// TIA Portal project "EbAndon v2_0_1" (V15) (continued)
TYPE "Color Library"
   STRUCT
      BkBk : USInt := 0;
      BgWh : USInt := 1;
      FgWh : USInt := 2;
      FlWh : USInt := 3;
      BgGray : USInt := 4;
      FgGray : USInt := 5;
      FlGray : USInt := 6;
      BgLRd : USInt := 7;
      FgLRd : USInt := 8;
      FlLRd : USInt := 9;
      BgDRd : USInt := 10;
      FgDRd : USInt := 11;
      FlDrd : USInt := 12;
      BgLYe : USInt := 13;
      FgLYe : USInt := 14;
      FlLYe : USInt := 15;
      BgDYe : USInt := 16;
      FgDYe : USInt := 17;
      FlDYe : USInt := 18;
      BgLGr : USInt := 19;
      FgLGr : USInt := 20;
      FlLGr : USInt := 21;
      BgDGr : USInt := 22;
      FgDGr : USInt := 23;
      FlDGr : USInt := 24;
      BgLTe : USInt := 25;
      FgLTe : USInt := 26;
      FlLTe : USInt := 27;
      BgDTe : USInt := 28;
      FgDTe : USInt := 29;
      FlDTe : USInt := 30;
      BgLBl : USInt := 31;
      FgLBl : USInt := 32;
      FlLBl : USInt := 33;
      BgDBl : USInt := 34;
      FgDBl : USInt := 35;
      FlDBl : USInt := 36;
      BgLPu : USInt := 37;
      FgLPu : USInt := 38;
      FlLPu : USInt := 39;
      BgDPu : USInt := 40;
      FgDPu : USInt := 41;
      FlDPu : USInt := 42;
      disabled : USInt := 254;
      invisible : USInt := 255;
   END_STRUCT;
END_TYPE

TYPE "Station Assignment: Button Details"
   STRUCT
      alloted : Struct
         animate : USInt;
         value : WString[10];
      END_STRUCT;
      critical : Struct
         animate : USInt;
         value : WString[10];
      END_STRUCT;
      label : Struct
         animate : USInt;
         value : WString[2];
      END_STRUCT;
      partNumber : Struct
         animate : USInt;
         value : WString[40];
      END_STRUCT;
      select : Struct
         actuate : Bool;
         animate : USInt;
      END_STRUCT;
   END_STRUCT;
END_TYPE

TYPE "IO Field Data: Part Number"
   STRUCT
      animate : USInt;
      inputFinished : Bool;
      value : WString[40];
   END_STRUCT;
END_TYPE

TYPE "Line Label Data"
   STRUCT
      animate : Struct
         bg : USInt;
         ioField : USInt;
      END_STRUCT;
      inputFinished : Bool;
      value : WString[10];
   END_STRUCT;
END_TYPE

TYPE "Drop Zone Data"
   STRUCT
      animate : Struct
         bg : USInt;
         ioField : USInt;
      END_STRUCT;
      inputFinished : Bool;
      value : WString[10];
   END_STRUCT;
END_TYPE

TYPE "IO Field Data: Timers"
   STRUCT
      animate : USInt;
      inputFinished : Bool;
      value : WString[5];
   END_STRUCT;
END_TYPE

TYPE "Table Nav"
   STRUCT
      top : "PB Data: Graphic/Text List";
      pageUp : "PB Data: Graphic/Text List";
      lineUp : "PB Data: Graphic/Text List";
      lineDown : "PB Data: Graphic/Text List";
      pageDown : "PB Data: Graphic/Text List";
      bottom : "PB Data: Graphic/Text List";
   END_STRUCT;
END_TYPE

DATA_BLOCK "EMP IDB"   // DB1
{ S7_Optimized_Access := 'TRUE' }
VERSION : 0.1
// stored: InstanceOfName EMP
"EMP"
BEGIN
   constants.buttonCount := 8;
   stations.current[0].presetTime.allotted[7] := 1800.0;
   stations.current[0].presetTime.allotted[3] := 1800.0;
   stations.current[0].presetTime.critical[7] := 300.0;
   stations.current[0].presetTime.critical[3] := 300.0;
   stations.current[0].partNumbers[7] := WSTRING#'16.32.112.500.100A';
   stations.current[0].partNumbers[6] := WSTRING#'';
   stations.current[0].partNumbers[5] := WSTRING#'';
   stations.current[0].partNumbers[3] := WSTRING#'16.32.112.500.220A';
   stations.current[0].partNumbers[2] := WSTRING#'';
   stations.current[0].partNumbers[1] := WSTRING#'';
   stations.current[0].line := WSTRING#'VOLVO 16';
   stations.current[1].line := WSTRING#'VOLVO 16';
   stations.current[2].line := WSTRING#'VOLVO 16';
   stations.current[0].dropZone := 1;
   stations.current[1].dropZone := 2;
   stations.current[2].dropZone := 3;
   stations.current[3].dropZone := 4;
   stations.current[3].line := WSTRING#'VOLVO 16';
   stations.current[4].dropZone := 5;
   stations.current[4].line := WSTRING#'VOLVO 16';
   stations.current[5].line := WSTRING#'VOLVO 16';
   stations.current[5].dropZone := 6;
   stations.current[6].dropZone := 7;
   stations.current[6].line := WSTRING#'VOLVO 16';
   stations.current[7].dropZone := 8;
   stations.current[7].line := WSTRING#'VOLVO 16';
   stations.current[8].dropZone := 9;
   stations.current[8].line := WSTRING#'VOLVO 16';
   stations.current[9].dropZone := 10;
   stations.current[9].line := WSTRING#'VOLVO 16';
   stations.current[10].dropZone := 11;
   stations.current[10].line := WSTRING#'VOLVO 16';
   stations.current[11].line := WSTRING#'CHM';
   stations.current[11].dropZone := 1;
   stations.current[12].line := WSTRING#'CHM';
   stations.current[12].dropZone := 2;
   stations.current[13].line := WSTRING#'CHM';
   stations.current[13].dropZone := 3;
   stations.current[14].dropZone := 4;
   stations.current[14].line := WSTRING#'CHM';
   stations.current[15].line := WSTRING#'CHM';
   stations.current[15].dropZone := 5;
   stations.current[16].dropZone := 1;
   stations.current[16].line := WSTRING#'CDO';
   stations.current[17].dropZone := 2;
   stations.current[17].line := WSTRING#'CDO';
   stations.current[18].line := WSTRING#'CDO';
   stations.current[18].dropZone := 3;
   stations.current[19].dropZone := 1;
   stations.current[19].line := WSTRING#'BFL';
   stations.current[20].dropZone := 2;
   stations.current[20].line := WSTRING#'BFL';
   stations.current[21].line := WSTRING#'BFL';
   stations.current[21].dropZone := 3;
   stations.current[22].dropZone := 1;
   stations.current[22].line := WSTRING#'LGS';
   stations.current[22].partNumbers[7] := WSTRING#'16.08.216.161.020A';
   stations.current[21].partNumbers[5] := WSTRING#'';
   stations.current[21].partNumbers[6] := WSTRING#'';
   stations.current[21].partNumbers[7] := WSTRING#'16.08.208.011.010G';
   stations.current[18].partNumbers[3] := WSTRING#'16.08.216.911.040B$L16.08.216.200.050A';
   stations.current[18].partNumbers[4] := WSTRING#'';
   stations.current[18].partNumbers[5] := WSTRING#'';
   stations.current[18].partNumbers[6] := WSTRING#'16.08.216.181.020A$L16.08.208.331.000F';
   stations.current[18].partNumbers[7] := WSTRING#'16.08.216.951.010A';
   stations.current[19].partNumbers[7] := WSTRING#'16.08.211.511.020F';
   stations.current[11].partNumbers[0] := WSTRING#'';
   stations.current[11].partNumbers[1] := WSTRING#'';
   stations.current[11].partNumbers[2] := WSTRING#'';
   stations.current[11].partNumbers[3] := WSTRING#'16.08.216.515.008C';
   stations.current[11].partNumbers[4] := WSTRING#'';
   stations.current[11].partNumbers[5] := WSTRING#'';
   stations.current[11].partNumbers[6] := WSTRING#'';
   stations.current[11].partNumbers[7] := WSTRING#'16.08.208.131.010L';
   stations.current[13].partNumbers[0] := WSTRING#'';
   stations.current[13].partNumbers[1] := WSTRING#'';
   stations.current[13].partNumbers[2] := WSTRING#'16.08.216.251.000B';
   stations.current[13].partNumbers[3] := WSTRING#'16.08.216.911.000G';
   stations.current[13].partNumbers[4] := WSTRING#'';
   stations.current[13].partNumbers[5] := WSTRING#'';
   stations.current[13].partNumbers[6] := WSTRING#'16.08.216.911.000H';
   stations.current[13].partNumbers[7] := WSTRING#'16.08.216.911.000C';
   stations.current[14].partNumbers[0] := WSTRING#'';
   stations.current[14].partNumbers[1] := WSTRING#'';
   stations.current[14].partNumbers[2] := WSTRING#'16.08.216.181.100A';
   stations.current[14].partNumbers[3] := WSTRING#'16.08.216.910.020B';
   stations.current[14].partNumbers[4] := WSTRING#'';
   stations.current[14].partNumbers[5] := WSTRING#'16.08.216.181.090A';
   stations.current[14].partNumbers[6] := WSTRING#'16.08.216.722.001A';
   stations.current[14].partNumbers[7] := WSTRING#'16.08.216.181.010B';
   stations.current[18].partNumbers[0] := WSTRING#'';
   stations.current[18].partNumbers[1] := WSTRING#'';
   stations.current[18].partNumbers[2] := WSTRING#'';
   stations.current[12].partNumbers[0] := WSTRING#'';
   stations.current[12].partNumbers[1] := WSTRING#'16.08.216.526.009A';
   stations.current[12].partNumbers[2] := WSTRING#'16.08.216.871.010C';
   stations.current[12].partNumbers[3] := WSTRING#'16.08.216.141.010C';
   stations.current[12].partNumbers[4] := WSTRING#'';
   stations.current[12].partNumbers[5] := WSTRING#'16.08.216.526.002C';
   stations.current[12].partNumbers[6] := WSTRING#'16.08.215.871.010C';
   stations.current[12].partNumbers[7] := WSTRING#'16.08.215.141.010C';
   stations.current[17].partNumbers[0] := WSTRING#'';
   stations.current[17].partNumbers[1] := WSTRING#'';
   stations.current[17].partNumbers[2] := WSTRING#'16.08.216.501.010A';
   stations.current[17].partNumbers[3] := WSTRING#'16.08.208.691.010D';
   stations.current[17].partNumbers[4] := WSTRING#'';
   stations.current[17].partNumbers[5] := WSTRING#'';
   stations.current[17].partNumbers[6] := WSTRING#'16.08.216.790.001A';
   stations.current[17].partNumbers[7] := WSTRING#'16.08.208.531.020L';
   stations.current[15].partNumbers[0] := WSTRING#'';
   stations.current[15].partNumbers[1] := WSTRING#'';
   stations.current[15].partNumbers[2] := WSTRING#'16.08.216.511.000C';
   stations.current[15].partNumbers[3] := WSTRING#'16.08.208.501.000B';
   stations.current[15].partNumbers[4] := WSTRING#'';
   stations.current[15].partNumbers[5] := WSTRING#'16.08.216.551.000B';
   stations.current[15].partNumbers[6] := WSTRING#'16.08.216.231.000B';
   stations.current[15].partNumbers[7] := WSTRING#'16.08.216.501.000C';
   stations.current[16].partNumbers[0] := WSTRING#'';
   stations.current[16].partNumbers[1] := WSTRING#'';
   stations.current[16].partNumbers[2] := WSTRING#'';
   stations.current[16].partNumbers[3] := WSTRING#'16.08.216.912.060B$L16.08.216.202.080A';
   stations.current[16].partNumbers[4] := WSTRING#'';
   stations.current[16].partNumbers[5] := WSTRING#'';
   stations.current[16].partNumbers[6] := WSTRING#'16.08.216.911.030B';
   stations.current[16].partNumbers[7] := WSTRING#'16.08.216.912.050A';
   stations.current[21].partNumbers[0] := WSTRING#'';
   stations.current[21].partNumbers[1] := WSTRING#'';
   stations.current[21].partNumbers[2] := WSTRING#'';
   stations.current[21].partNumbers[3] := WSTRING#'';
   stations.current[21].partNumbers[4] := WSTRING#'';
   stations.current[20].partNumbers[0] := WSTRING#'';
   stations.current[20].partNumbers[1] := WSTRING#'';
   stations.current[20].partNumbers[2] := WSTRING#'';
   stations.current[20].partNumbers[3] := WSTRING#'';
   stations.current[20].partNumbers[4] := WSTRING#'';
   stations.current[20].partNumbers[5] := WSTRING#'';
   stations.current[20].partNumbers[6] := WSTRING#'';
   stations.current[20].partNumbers[7] := WSTRING#'PEANUTS';
   stations.current[8].partNumbers[0] := WSTRING#'';
   stations.current[8].partNumbers[1] := WSTRING#'';
   stations.current[8].partNumbers[2] := WSTRING#'';
   stations.current[8].partNumbers[3] := WSTRING#'16.32.112.580.020A';
   stations.current[8].partNumbers[4] := WSTRING#'';
   stations.current[8].partNumbers[5] := WSTRING#'';
   stations.current[8].partNumbers[6] := WSTRING#'16.32.112.500.300E';
   stations.current[8].partNumbers[7] := WSTRING#'16.32.112.520.300E';
   stations.current[9].partNumbers[0] := WSTRING#'';
   stations.current[9].partNumbers[1] := WSTRING#'';
   stations.current[9].partNumbers[2] := WSTRING#'';
   stations.current[9].partNumbers[3] := WSTRING#'16.32.112.594.000C';
   stations.current[9].partNumbers[4] := WSTRING#'';
   stations.current[9].partNumbers[5] := WSTRING#'';
   stations.current[9].partNumbers[6] := WSTRING#'';
   stations.current[9].partNumbers[7] := WSTRING#'16.32.112.584.000C';
   stations.current[10].partNumbers[0] := WSTRING#'';
   stations.current[10].partNumbers[1] := WSTRING#'';
   stations.current[10].partNumbers[2] := WSTRING#'';
   stations.current[10].partNumbers[3] := WSTRING#'16.32.112.500.150B';
   stations.current[10].partNumbers[4] := WSTRING#'';
   stations.current[10].partNumbers[5] := WSTRING#'';
   stations.current[10].partNumbers[6] := WSTRING#'16.32.806.502.080A';
   stations.current[10].partNumbers[7] := WSTRING#'16.32.112.500.160A';
   stations.current[0].partNumbers[0] := WSTRING#'';
   stations.current[0].partNumbers[4] := WSTRING#'';
   stations.current[1].partNumbers[0] := WSTRING#'';
   stations.current[1].partNumbers[1] := WSTRING#'';
   stations.current[1].partNumbers[2] := WSTRING#'16.32.112.509.070A';
   stations.current[1].partNumbers[3] := WSTRING#'16.32.112.704.000C';
   stations.current[1].partNumbers[4] := WSTRING#'';
   stations.current[1].partNumbers[5] := WSTRING#'';
   stations.current[1].partNumbers[6] := WSTRING#'16.32.112.504.060A';
   stations.current[1].partNumbers[7] := WSTRING#'16.32.112.500.060D';
   stations.current[2].partNumbers[0] := WSTRING#'';
   stations.current[2].partNumbers[1] := WSTRING#'16.32.112.509.050E';
   stations.current[2].partNumbers[2] := WSTRING#'16.32.112.504.070G';
   stations.current[2].partNumbers[3] := WSTRING#'16.32.112.851.001A';
   stations.current[2].partNumbers[4] := WSTRING#'';
   stations.current[2].partNumbers[5] := WSTRING#'16.32.112.509.080F';
   stations.current[2].partNumbers[6] := WSTRING#'16.32.112.870.000C';
   stations.current[2].partNumbers[7] := WSTRING#'16.32.112.851.000A';
   stations.current[3].partNumbers[0] := WSTRING#'';
   stations.current[3].partNumbers[1] := WSTRING#'16.32.112.522.130A';
   stations.current[3].partNumbers[2] := WSTRING#'16.32.112.522.050A';
   stations.current[3].partNumbers[3] := WSTRING#'16.32.112.521.020B';
   stations.current[3].partNumbers[4] := WSTRING#'';
   stations.current[3].partNumbers[5] := WSTRING#'16.32.112.522.040D';
   stations.current[3].partNumbers[6] := WSTRING#'16.32.112.521.010B';
   stations.current[3].partNumbers[7] := WSTRING#'16.32.112.521.030A';
   stations.current[4].partNumbers[0] := WSTRING#'';
   stations.current[4].partNumbers[1] := WSTRING#'';
   stations.current[4].partNumbers[2] := WSTRING#'';
   stations.current[4].partNumbers[3] := WSTRING#'';
   stations.current[4].partNumbers[4] := WSTRING#'';
   stations.current[4].partNumbers[5] := WSTRING#'';
   stations.current[4].partNumbers[6] := WSTRING#'';
   stations.current[4].partNumbers[7] := WSTRING#'16.32.112.529.020B';
   stations.current[5].partNumbers[0] := WSTRING#'';
   stations.current[5].partNumbers[1] := WSTRING#'16.32.112.529.010A';
   stations.current[5].partNumbers[2] := WSTRING#'16.32.112.529.030A';
   stations.current[5].partNumbers[3] := WSTRING#'16.32.112.502.060B';
   stations.current[5].partNumbers[4] := WSTRING#'';
   stations.current[5].partNumbers[5] := WSTRING#'16.32.112.529.050D';
   stations.current[5].partNumbers[6] := WSTRING#'16.32.112.502.070E';
   stations.current[5].partNumbers[7] := WSTRING#'16.32.112.502.050B';
   stations.current[6].partNumbers[0] := WSTRING#'';
   stations.current[6].partNumbers[1] := WSTRING#'16.32.112.621.020A';
   stations.current[6].partNumbers[2] := WSTRING#'16.32.112.621.010A';
   stations.current[6].partNumbers[3] := WSTRING#'16.32.112.751.000D';
   stations.current[6].partNumbers[4] := WSTRING#'';
   stations.current[6].partNumbers[5] := WSTRING#'16.32.112.751.001C';
   stations.current[6].partNumbers[6] := WSTRING#'16.32.112.601.040A';
   stations.current[6].partNumbers[7] := WSTRING#'16.32.112.601.030A';
   stations.current[7].partNumbers[0] := WSTRING#'';
   stations.current[7].partNumbers[1] := WSTRING#'';
   stations.current[7].partNumbers[2] := WSTRING#'';
   stations.current[7].partNumbers[3] := WSTRING#'16.32.112.500.520B';
   stations.current[7].partNumbers[4] := WSTRING#'';
   stations.current[7].partNumbers[5] := WSTRING#'';
   stations.current[7].partNumbers[6] := WSTRING#'16.32.112.500.090B';
   stations.current[7].partNumbers[7] := WSTRING#'16.32.112.500.120A';
   stations.current[23].line := WSTRING#'LGS';
   stations.current[23].dropZone := 2;
   stations.current[23].partNumbers[0] := WSTRING#'';
   stations.current[23].partNumbers[1] := WSTRING#'';
   stations.current[23].partNumbers[2] := WSTRING#'';
   stations.current[23].partNumbers[3] := WSTRING#'';
   stations.current[23].partNumbers[4] := WSTRING#'';
   stations.current[23].partNumbers[5] := WSTRING#'';
   stations.current[23].partNumbers[6] := WSTRING#'';
   stations.current[23].partNumbers[7] := WSTRING#'16.08.208.021.020C';
   stations.current[22].partNumbers[0] := WSTRING#'';
   stations.current[22].partNumbers[1] := WSTRING#'';
   stations.current[22].partNumbers[2] := WSTRING#'';
   stations.current[22].partNumbers[3] := WSTRING#'16.08.208.161.020F';
   stations.current[22].partNumbers[4] := WSTRING#'';
   stations.current[22].partNumbers[5] := WSTRING#'';
   stations.current[22].partNumbers[6] := WSTRING#'OP60 - STAMPINGS';
   stations.current[19].partNumbers[0] := WSTRING#'';
   stations.current[19].partNumbers[1] := WSTRING#'';
   stations.current[19].partNumbers[2] := WSTRING#'16.08.216.831.020A';
   stations.current[19].partNumbers[3] := WSTRING#'16.08.208.151.010F';
   stations.current[19].partNumbers[4] := WSTRING#'';
   stations.current[19].partNumbers[5] := WSTRING#'16.08.217.411.080A';
   stations.current[19].partNumbers[6] := WSTRING#'16.08.216.151.010B';
   constants.hmiRowCount := 12;
   constants.ledRowCount := 12;
END_DATA_BLOCK

DATA_BLOCK "HMI"   // DB2
{ S7_Optimized_Access := 'TRUE' }
VERSION : 0.1
   VAR
      partCall : "Part Call Screen";
      screenNumber : Int;
      settings : "Settings Screen";
      barcode : "Barcode Screen";
      tableNav : "Table Nav";
   END_VAR
BEGIN
   settings.current.kp8.buttons[1].label := WSTRING#'6';
   settings.current.kp8.buttons[2].label := WSTRING#'4';
   settings.current.kp8.buttons[3].label := WSTRING#'2';
   settings.current.kp8.buttons[5].label := WSTRING#'5';
   settings.current.kp8.buttons[6].label := WSTRING#'3';
   settings.current.kp8.buttons[7].label := WSTRING#'1';
END_DATA_BLOCK

DATA_BLOCK "Parts"   // DB3
{ S7_Optimized_Access := 'TRUE' }
VERSION : 0.1
   VAR
      pRow : Int;
   END_VAR
   VAR RETAIN
      requests : "Part Request Data";
   END_VAR
BEGIN
END_DATA_BLOCK

DATA_BLOCK "LED Sign"   // DB4
{ S7_Optimized_Access := 'TRUE' }
VERSION : 0.1
   VAR
      request : "LED Sign Data";
   END_VAR
BEGIN
END_DATA_BLOCK

FUNCTION_BLOCK "EMP"   // FB1, LAD
{ S7_Optimized_Access := 'TRUE' }
VERSION : 0.1
   VAR RETAIN
      constants : "Constants";
   END_VAR
   VAR
      instBaseAnimations : "Base Animations";
      instHMIAnimations : "Format Part Call Requests";
      instInitialize : "Initialize";
      instKP8ButtonActivation : "KP8 Button Activation";
      instKP8ExpandedAnimations : "KP8 Expanded Animations";
      instPartTimers : "Part Timers";
      instRecordPartRequest : "Record Part Request";
      instRemovePartRequest : "Remove Part Request";
      instResetInitRequest : "Reset Init Requests";
      instStackLightAnimations : "Stack Light Animations";
      "KP8 Drivers" : Array[0..#stationCount] of "KP8 Driver";
   END_VAR
   VAR RETAIN
      stations : "Stations";
   END_VAR
   VAR
      instHMIBarcode : "HMI Barcod Screen";
      instCollapseTable : "Collapse Table";
      instPopulateHMI : "HMI Populate Part Call";
      instHMISettings : "HMI Settings Screen";
      instClearReqData : "Clear Part Requests";
      instDefaultTmrPrst : "Load Default Timer Presets";
      instPopulateLED : "LED Populate Sign";
   END_VAR
   VAR_TEMP
      i : Int;
      stnCount : Int;
   END_VAR
   VAR CONSTANT
      stationCount : Int := 24;
   END_VAR
BEGIN

REGION Network 1: PHYSICAL TO GLOBAL
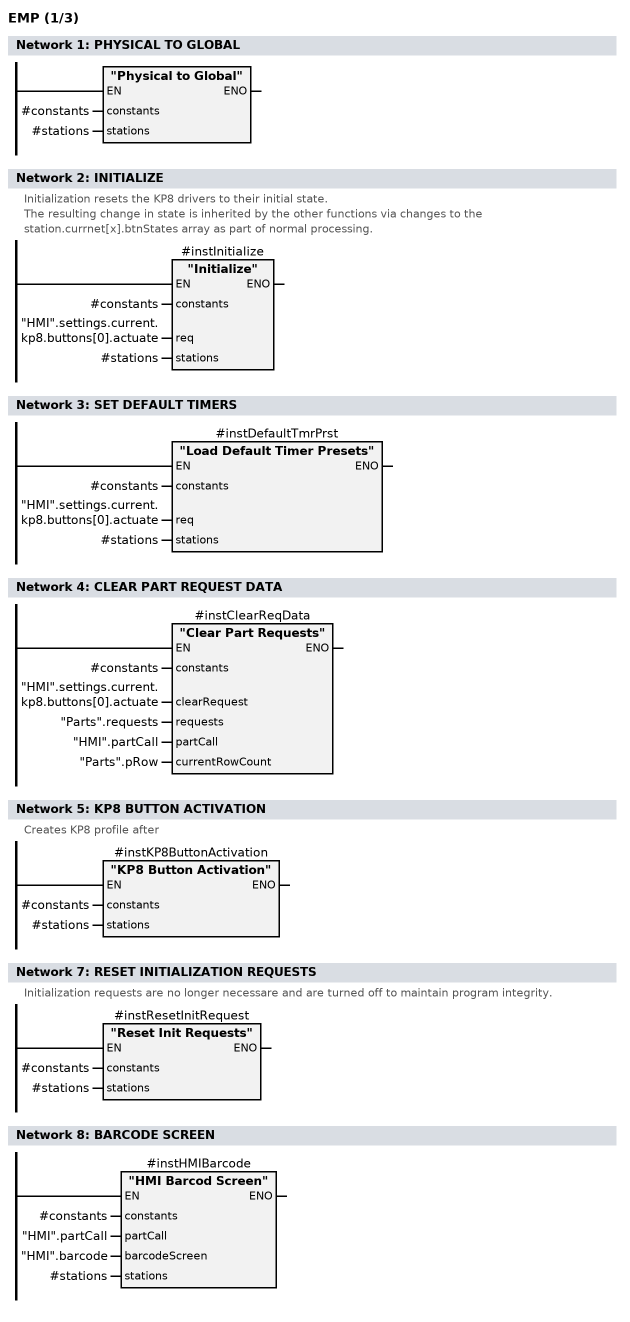
   RUNG wire#powerrail
      "Physical to Global"(constants := #constants, stations := #stations)
   END_RUNG
   // the same network as SCL:
   "Physical to Global"(constants := #constants, stations := #stations);
END_REGION

REGION Network 2: INITIALIZE
   // Initialization resets the KP8 drivers to their initial state.
   // The resulting change in state is inherited by the other functions via changes to the
   // station.currnet[x].btnStates array as part of normal processing.
   RUNG wire#powerrail
      #instInitialize(constants := #constants, req := "HMI".settings.current.kp8.buttons[0].actuate, stations := #stations)
   END_RUNG
   // the same network as SCL:
   #instInitialize(constants := #constants,   // "Initialize"
                   req := "HMI".settings.current.kp8.buttons[0].actuate,
                   stations := #stations);
END_REGION

REGION Network 3: SET DEFAULT TIMERS
   RUNG wire#powerrail
      #instDefaultTmrPrst(constants := #constants, req := "HMI".settings.current.kp8.buttons[0].actuate, stations := #stations)
   END_RUNG
   // the same network as SCL:
   #instDefaultTmrPrst(constants := #constants,   // "Load Default Timer Presets"
                       req := "HMI".settings.current.kp8.buttons[0].actuate,
                       stations := #stations);
END_REGION

REGION Network 4: CLEAR PART REQUEST DATA
   RUNG wire#powerrail
      #instClearReqData(constants := #constants, clearRequest := "HMI".settings.current.kp8.buttons[0].actuate, requests := "Parts".requests, partCall := "HMI".partCall, currentRowCount := "Parts".pRow)
   END_RUNG
   // the same network as SCL:
   #instClearReqData(constants := #constants,   // "Clear Part Requests"
                     clearRequest := "HMI".settings.current.kp8.buttons[0].actuate,
                     requests := "Parts".requests,
                     partCall := "HMI".partCall,
                     currentRowCount := "Parts".pRow);
END_REGION

REGION Network 5: KP8 BUTTON ACTIVATION
   // Creates KP8 profile after
   RUNG wire#powerrail
      #instKP8ButtonActivation(constants := #constants, stations := #stations)
   END_RUNG
   // the same network as SCL:
   #instKP8ButtonActivation(constants := #constants, stations := #stations);   // "KP8 Button Activation"
END_REGION

REGION Network 6 (SCL): KP8 DRIVER CALLS
   REGION "LOOP THROUGH STATIONS"
       #stnCount := #constants.stationCount - 1;
       FOR #i := 0 TO #stnCount DO
           #"KP8 Drivers"[#i](btnIn := #stations.current[#i].kp8In,
                              hardInit := #stations.current[#i].init.hard,
                              softInit := #stations.current[#i].init.soft,
                              btn0Activate := #stations.current[#i].kp8Config.activate[0],
                              btn0Mode := #stations.current[#i].kp8Config.mode[0],
                              btn0Group := #stations.current[#i].kp8Config.group[0],
                              btn0Flash := #stations.current[#i].kp8Config.flash[0],
                              btn0ColorOn1 := #stations.current[#i].kp8Config.colorOn1[0],
                              btn0ColorOn2 := #stations.current[#i].kp8Config.colorOn2[0],
                              btn0ColorOff := #stations.current[#i].kp8Config.colorOff[0],
                              btn1Activate := #stations.current[#i].kp8Config.activate[1],
                              btn1Mode := #stations.current[#i].kp8Config.mode[1],
                              btn1Group := #stations.current[#i].kp8Config.group[1],
                              btn1Flash := #stations.current[#i].kp8Config.flash[1],
                              btn1ColorOn1 := #stations.current[#i].kp8Config.colorOn1[1],
                              btn1ColorOn2 := #stations.current[#i].kp8Config.colorOn2[1],
                              btn1ColorOff := #stations.current[#i].kp8Config.colorOff[1],
                              btn2Activate := #stations.current[#i].kp8Config.activate[2],
                              btn2Mode := #stations.current[#i].kp8Config.mode[2],
                              btn2Group := #stations.current[#i].kp8Config.group[2],
                              btn2Flash := #stations.current[#i].kp8Config.flash[2],
                              btn2ColorOn1 := #stations.current[#i].kp8Config.colorOn1[2],
                              btn2ColorOn2 := #stations.current[#i].kp8Config.colorOn2[2],
                              btn2ColorOff := #stations.current[#i].kp8Config.colorOff[2],
                              btn3Activate := #stations.current[#i].kp8Config.activate[3],
                              btn3Mode := #stations.current[#i].kp8Config.mode[3],
                              btn3Group := #stations.current[#i].kp8Config.group[3],
                              btn3Flash := #stations.current[#i].kp8Config.flash[3],
                              btn3ColorOn1 := #stations.current[#i].kp8Config.colorOn1[3],
                              btn3ColorOn2 := #stations.current[#i].kp8Config.colorOn2[3],
                              btn3ColorOff := #stations.current[#i].kp8Config.colorOff[3],
                              btn4Activate := #stations.current[#i].kp8Config.activate[4],
                              btn4Mode := #stations.current[#i].kp8Config.mode[4],
                              btn4Group := #stations.current[#i].kp8Config.group[4],
                              btn4Flash := #stations.current[#i].kp8Config.flash[4],
                              btn4ColorOn1 := #stations.current[#i].kp8Config.colorOn1[4],
                              btn4ColorOn2 := #stations.current[#i].kp8Config.colorOn2[4],
                              btn4ColorOff := #stations.current[#i].kp8Config.colorOff[4],
                              btn5Activate := #stations.current[#i].kp8Config.activate[5],
                              btn5Mode := #stations.current[#i].kp8Config.mode[5],
                              btn5Group := #stations.current[#i].kp8Config.group[5],
                              btn5Flash := #stations.current[#i].kp8Config.flash[5],
                              btn5ColorOn1 := #stations.current[#i].kp8Config.colorOn1[5],
                              btn5ColorOn2 := #stations.current[#i].kp8Config.colorOn2[5],
                              btn5ColorOff := #stations.current[#i].kp8Config.colorOff[5],
                              btn6Activate := #stations.current[#i].kp8Config.activate[6],
                              btn6Mode := #stations.current[#i].kp8Config.mode[6],
                              btn6Group := #stations.current[#i].kp8Config.group[6],
                              btn6Flash := #stations.current[#i].kp8Config.flash[6],
                              btn6ColorOn1 := #stations.current[#i].kp8Config.colorOn1[6],
                              btn6ColorOn2 := #stations.current[#i].kp8Config.colorOn2[6],
                              btn6ColorOff := #stations.current[#i].kp8Config.colorOff[6],
                              btn7Activate := #stations.current[#i].kp8Config.activate[7],
                              btn7Mode := #stations.current[#i].kp8Config.mode[7],
                              btn7Group := #stations.current[#i].kp8Config.group[7],
                              btn7Flash := #stations.current[#i].kp8Config.flash[7],
                              btn7ColorOn1 := #stations.current[#i].kp8Config.colorOn1[7],
                              btn7ColorOn2 := #stations.current[#i].kp8Config.colorOn2[7],
                              btn7ColorOff := #stations.current[#i].kp8Config.colorOff[7],
                              btnStatesOut => #stations.current[#i].btnStates,
                              btnColorsOut => #stations.current[#i].kp8Out);
       END_FOR;
   END_REGION
END_REGION

REGION Network 7: RESET INITIALIZATION REQUESTS
   // Initialization requests are no longer necessare and are turned off to maintain program integrity.
   RUNG wire#powerrail
      #instResetInitRequest(constants := #constants, stations := #stations)
   END_RUNG
   // the same network as SCL:
   #instResetInitRequest(constants := #constants, stations := #stations);   // "Reset Init Requests"
END_REGION

REGION Network 8: BARCODE SCREEN
   RUNG wire#powerrail
      #instHMIBarcode(constants := #constants, partCall := "HMI".partCall, barcodeScreen := "HMI".barcode, stations := #stations)
   END_RUNG
   // the same network as SCL:
   #instHMIBarcode(constants := #constants,   // "HMI Barcod Screen"
                   partCall := "HMI".partCall,
                   barcodeScreen := "HMI".barcode,
                   stations := #stations);
END_REGION

REGION Network 9: PART TIMERS
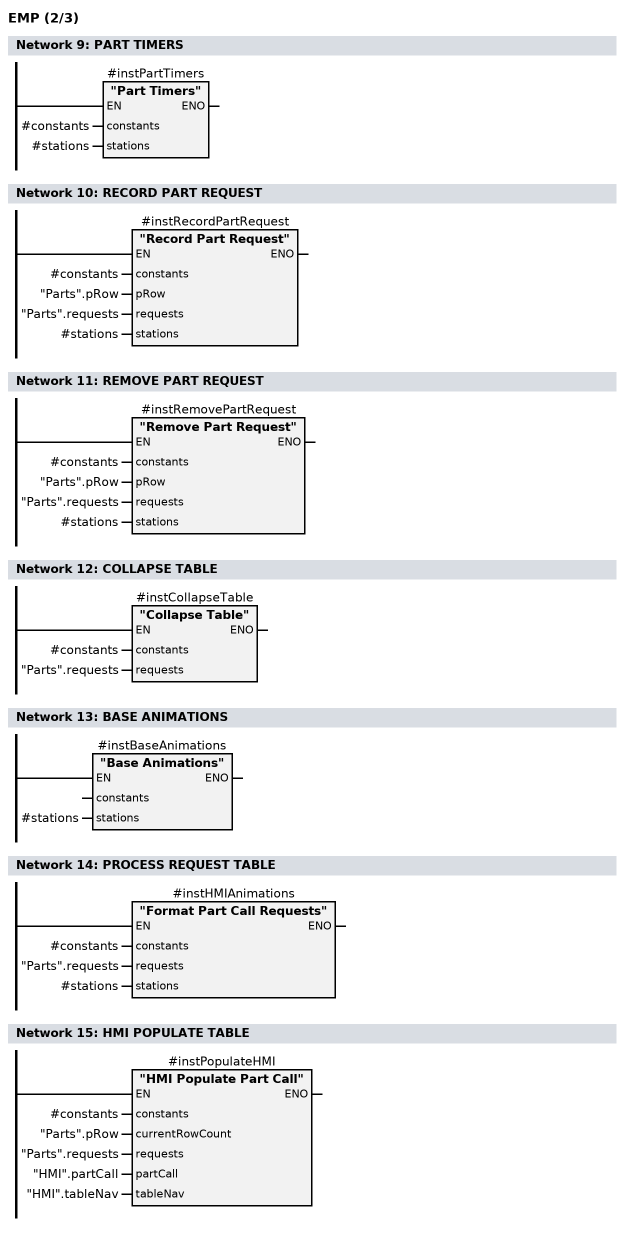
   RUNG wire#powerrail
      #instPartTimers(constants := #constants, stations := #stations)
   END_RUNG
   // the same network as SCL:
   #instPartTimers(constants := #constants, stations := #stations);   // "Part Timers"
END_REGION

REGION Network 10: RECORD PART REQUEST
   RUNG wire#powerrail
      #instRecordPartRequest(constants := #constants, pRow := "Parts".pRow, requests := "Parts".requests, stations := #stations)
   END_RUNG
   // the same network as SCL:
   #instRecordPartRequest(constants := #constants,   // "Record Part Request"
                          pRow := "Parts".pRow,
                          requests := "Parts".requests,
                          stations := #stations);
END_REGION

REGION Network 11: REMOVE PART REQUEST
   RUNG wire#powerrail
      #instRemovePartRequest(constants := #constants, pRow := "Parts".pRow, requests := "Parts".requests, stations := #stations)
   END_RUNG
   // the same network as SCL:
   #instRemovePartRequest(constants := #constants,   // "Remove Part Request"
                          pRow := "Parts".pRow,
                          requests := "Parts".requests,
                          stations := #stations);
END_REGION

REGION Network 12: COLLAPSE TABLE
   RUNG wire#powerrail
      #instCollapseTable(constants := #constants, requests := "Parts".requests)
   END_RUNG
   // the same network as SCL:
   #instCollapseTable(constants := #constants, requests := "Parts".requests);   // "Collapse Table"
END_REGION

REGION Network 13: BASE ANIMATIONS
   RUNG wire#powerrail
      #instBaseAnimations(constants :=, stations := #stations)
   END_RUNG
   // the same network as SCL:
   #instBaseAnimations(stations := #stations);   // "Base Animations"
END_REGION

REGION Network 14: PROCESS REQUEST TABLE
   RUNG wire#powerrail
      #instHMIAnimations(constants := #constants, requests := "Parts".requests, stations := #stations)
   END_RUNG
   // the same network as SCL:
   #instHMIAnimations(constants := #constants, requests := "Parts".requests, stations := #stations);   // "Format Part Call Requests"
END_REGION
